   IF #_w2 THEN "DB_GlobalData".AKD.AKD1.wNewJobNumber := 4; END_IF;
   "reserve(3)":P := #_w2 AND NOT "reserve(2)";
END_REGION

REGION Network 5
   RUNG wire#powerrail
      Contact( "Clock_5Hz" )
      Coil( "xActuatorStatus" )
   END_RUNG
   // the same network as SCL:
   "xActuatorStatus" := "Clock_5Hz";
END_REGION

REGION Network 6
   #_w1 := "i_xSystemTrigger":P AND NOT "p_trig_trigg";   // rising edge
   "p_trig_trigg" := "i_xSystemTrigger":P;
   "r_eege_triger" := #_w1;
   "DB_safetyActuator".On_timer[1].TON(IN := "reserve(2)", PT := T#700ms);
END_REGION

REGION Network 7 (SCL)
   IF "r_eege_triger" THEN
       "tooglebit" := NOT "tooglebit";
   END_IF;
END_REGION

REGION Network 8
   RUNG wire#powerrail
      Contact( "DB_safetyActuator".On_timer[1].Q )
      R_Coil( "tooglebit" )
   END_RUNG
   // the same network as SCL:
   IF "DB_safetyActuator".On_timer[1].Q THEN "tooglebit" := FALSE; END_IF;
END_REGION

REGION Network 11: AKD1
   RUNG wire#powerrail
      Contact( "AKD_PNU_DATA".AKD1.PNU_userSETTINGS.xRadAKDTemp )
      Move(in := "AKD_PNU_DATA".AKD1.PNU_userSETTINGS.PNU_const.AKD_TEMP.PNU_number, out1 => "AKD_PNU_DATA".AKD1.PNU_DATA.to_PNU.iPNUnumber)
      Move(in := "AKD_PNU_DATA".AKD1.PNU_userSETTINGS.PNU_const.AKD_TEMP.PNU_subIndex, out1 => "AKD_PNU_DATA".AKD1.PNU_DATA.to_PNU.iPNUsubindex)
      Move(in := "AKD_PNU_DATA".AKD1.PNU_userSETTINGS.PNU_const.AKD_TEMP.PNU_type, out1 => "AKD_PNU_DATA".AKD1.PNU_DATA.to_PNU.wFormat)
      S_Coil( "AKD_PNU_DATA".AKD1.PNU_DATA.to_PNU.cmd.xStartRead )
      R_Coil( "AKD_PNU_DATA".AKD1.PNU_userSETTINGS.xRadAKDTemp )
   END_RUNG
   // the same network as SCL:
   IF "AKD_PNU_DATA".AKD1.PNU_userSETTINGS.xRadAKDTemp THEN
       "AKD_PNU_DATA".AKD1.PNU_DATA.to_PNU.iPNUnumber := "AKD_PNU_DATA".AKD1.PNU_userSETTINGS.PNU_const.AKD_TEMP.PNU_number;
       "AKD_PNU_DATA".AKD1.PNU_DATA.to_PNU.iPNUsubindex := "AKD_PNU_DATA".AKD1.PNU_userSETTINGS.PNU_const.AKD_TEMP.PNU_subIndex;
       "AKD_PNU_DATA".AKD1.PNU_DATA.to_PNU.wFormat := "AKD_PNU_DATA".AKD1.PNU_userSETTINGS.PNU_const.AKD_TEMP.PNU_type;
       "AKD_PNU_DATA".AKD1.PNU_DATA.to_PNU.cmd.xStartRead := TRUE;
       "AKD_PNU_DATA".AKD1.PNU_userSETTINGS.xRadAKDTemp := FALSE;
   END_IF;
END_REGION

REGION Network 12: read temperature every 0.5s
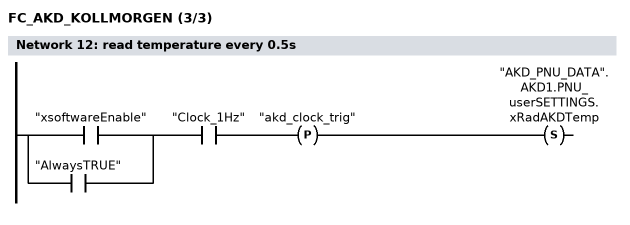
   RUNG wire#powerrail
      Contact( "xsoftwareEnable" )
      wire#w1
      Contact( "Clock_1Hz" )
      P_Trig( "akd_clock_trig" )
      S_Coil( "AKD_PNU_DATA".AKD1.PNU_userSETTINGS.xRadAKDTemp )
   END_RUNG
   RUNG wire#powerrail
      Contact( "AlwaysTRUE" )
   END_RUNG wire#w1
   // the same network as SCL:
   #_w1 := ("xsoftwareEnable" OR "AlwaysTRUE") AND "Clock_1Hz";
   #_w2 := #_w1 AND NOT "akd_clock_trig";   // rising edge
   "akd_clock_trig" := #_w1;
   IF #_w2 THEN "AKD_PNU_DATA".AKD1.PNU_userSETTINGS.xRadAKDTemp := TRUE; END_IF;
END_REGION
END_FUNCTION

FUNCTION "FC_RTD_DATA" : Void   // FC7, LAD
{ S7_Optimized_Access := 'TRUE' }
VERSION : 0.1
BEGIN

REGION Network 1
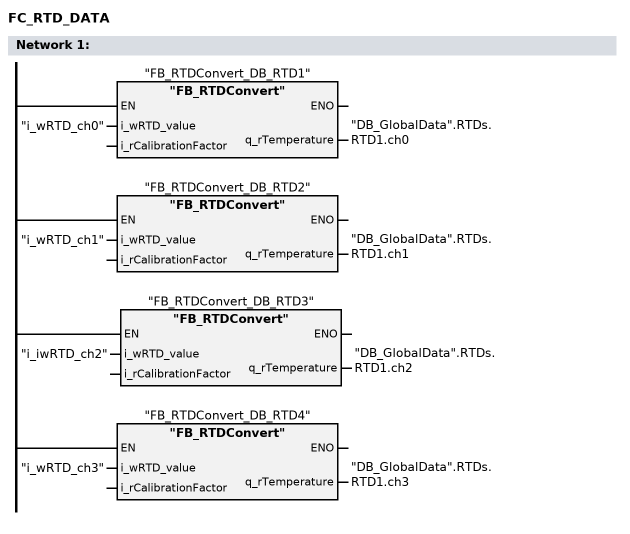
   RUNG wire#powerrail
      "FB_RTDConvert_DB_RTD1"(i_wRTD_value := "i_wRTD_ch0", i_rCalibrationFactor :=, q_rTemperature => "DB_GlobalData".RTDs.RTD1.ch0)
   END_RUNG
   RUNG wire#powerrail
      "FB_RTDConvert_DB_RTD2"(i_wRTD_value := "i_wRTD_ch1", i_rCalibrationFactor :=, q_rTemperature => "DB_GlobalData".RTDs.RTD1.ch1)
   END_RUNG
   RUNG wire#powerrail
      "FB_RTDConvert_DB_RTD3"(i_wRTD_value := "i_iwRTD_ch2", i_rCalibrationFactor :=, q_rTemperature => "DB_GlobalData".RTDs.RTD1.ch2)
   END_RUNG
   RUNG wire#powerrail
      "FB_RTDConvert_DB_RTD4"(i_wRTD_value := "i_wRTD_ch3", i_rCalibrationFactor :=, q_rTemperature => "DB_GlobalData".RTDs.RTD1.ch3)
   END_RUNG
   // the same network as SCL:
   "FB_RTDConvert_DB_RTD1"(i_wRTD_value := "i_wRTD_ch0", q_rTemperature => "DB_GlobalData".RTDs.RTD1.ch0);   // "FB_RTDConvert"
   "FB_RTDConvert_DB_RTD2"(i_wRTD_value := "i_wRTD_ch1", q_rTemperature => "DB_GlobalData".RTDs.RTD1.ch1);   // "FB_RTDConvert"
   "FB_RTDConvert_DB_RTD3"(i_wRTD_value := "i_iwRTD_ch2", q_rTemperature => "DB_GlobalData".RTDs.RTD1.ch2);   // "FB_RTDConvert"
   "FB_RTDConvert_DB_RTD4"(i_wRTD_value := "i_wRTD_ch3", q_rTemperature => "DB_GlobalData".RTDs.RTD1.ch3);   // "FB_RTDConvert"
END_REGION
END_FUNCTION

FUNCTION "FC_MQTT" : Void   // FC8, LAD
{ S7_Optimized_Access := 'TRUE' }
VERSION : 0.1
   VAR_TEMP
      globalstring : String;
      testbit : Bool;
   END_VAR
   VAR_TEMP   // added for the SCL form of the ladder/FBD networks
      _w1 : Bool;
   END_VAR
BEGIN

REGION Network 1
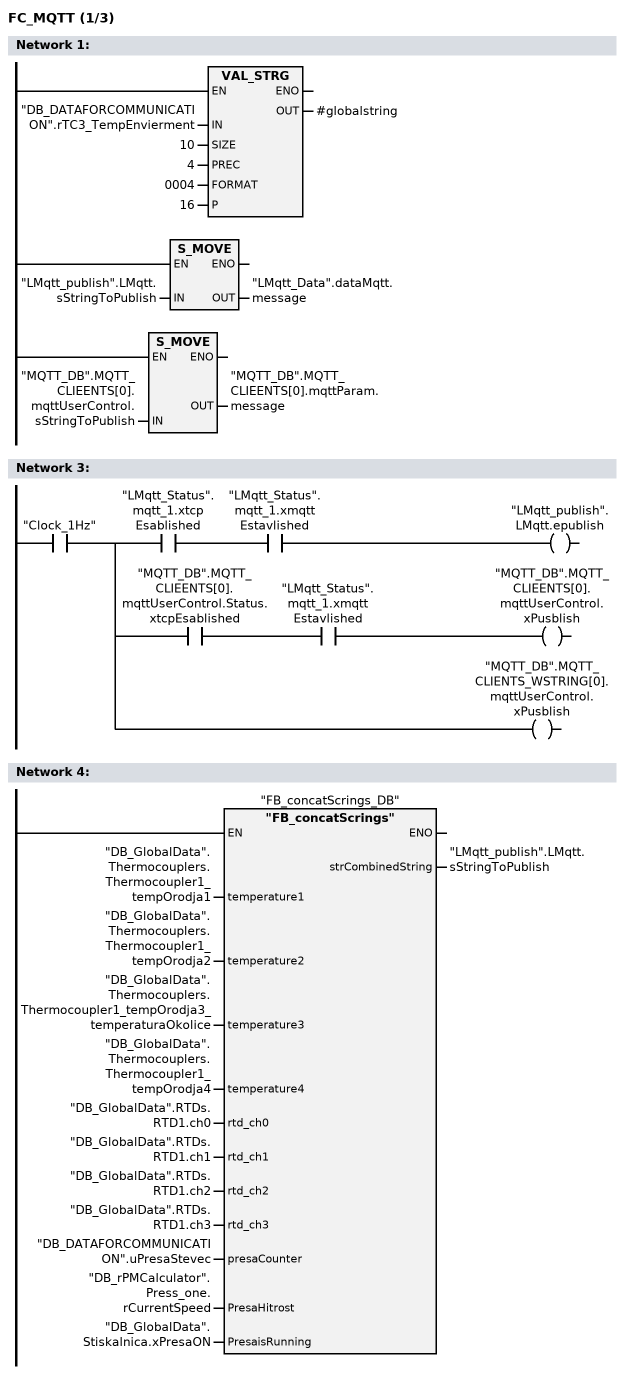
   VAL_STRG(IN := "DB_DATAFORCOMMUNICATION".rTC3_TempEnvierment,
            SIZE := 10,
            PREC := 4,
            FORMAT := 0004,
            P := 16,
            OUT => #globalstring);
   "LMqtt_Data".dataMqtt.message := "LMqtt_publish".LMqtt.sStringToPublish;
   "MQTT_DB".MQTT_CLIEENTS[0].mqttParam.message := "MQTT_DB".MQTT_CLIEENTS[0].mqttUserControl.sStringToPublish;
END_REGION

REGION Network 3
   RUNG wire#powerrail
      Contact( "Clock_1Hz" )
      wire#w1
      Contact( "LMqtt_Status".mqtt_1.xtcpEsablished )
      Contact( "LMqtt_Status".mqtt_1.xmqttEstavlished )
      Coil( "LMqtt_publish".LMqtt.epublish )
   END_RUNG
   RUNG wire#w1
      Contact( "MQTT_DB".MQTT_CLIEENTS[0].mqttUserControl.Status.xtcpEsablished )
      Contact( "LMqtt_Status".mqtt_1.xmqttEstavlished )
      Coil( "MQTT_DB".MQTT_CLIEENTS[0].mqttUserControl.xPusblish )
   END_RUNG
   RUNG wire#w1
      Coil( "MQTT_DB".MQTT_CLIENTS_WSTRING[0].mqttUserControl.xPusblish )
   END_RUNG
   // the same network as SCL:
   "LMqtt_publish".LMqtt.epublish := "Clock_1Hz" AND "LMqtt_Status".mqtt_1.xtcpEsablished AND "LMqtt_Status".mqtt_1.xmqttEstavlished;
   "MQTT_DB".MQTT_CLIEENTS[0].mqttUserControl.xPusblish := "Clock_1Hz" AND "MQTT_DB".MQTT_CLIEENTS[0].mqttUserControl.Status.xtcpEsablished AND "LMqtt_Status".mqtt_1.xmqttEstavlished;
   "MQTT_DB".MQTT_CLIENTS_WSTRING[0].mqttUserControl.xPusblish := "Clock_1Hz";
END_REGION

REGION Network 4
   RUNG wire#powerrail
      "FB_concatScrings_DB"(temperature1 := "DB_GlobalData".Thermocouplers.Thermocoupler1_tempOrodja1, temperature2 := "DB_GlobalData".Thermocouplers.Thermocoupler1_tempOrodja2, temperature3 := "DB_GlobalData".Thermocouplers.Thermocoupler1_tempOrodja3_temperaturaOkolice, temperature4 := "DB_GlobalData".Thermocouplers.Thermocoupler1_tempOrodja4, rtd_ch0 := "DB_GlobalData".RTDs.RTD1.ch0, rtd_ch1 := "DB_GlobalData".RTDs.RTD1.ch1, rtd_ch2 := "DB_GlobalData".RTDs.RTD1.ch2, rtd_ch3 := "DB_GlobalData".RTDs.RTD1.ch3, presaCounter := "DB_DATAFORCOMMUNICATION".uPresaStevec, PresaHitrost := "DB_rPMCalculator".Press_one.rCurrentSpeed, PresaisRunning := "DB_GlobalData".Stiskalnica.xPresaON, strCombinedString => "LMqtt_publish".LMqtt.sStringToPublish)
   END_RUNG
   // the same network as SCL:
   "FB_concatScrings_DB"(temperature1 := "DB_GlobalData".Thermocouplers.Thermocoupler1_tempOrodja1,   // "FB_concatScrings"
                         temperature2 := "DB_GlobalData".Thermocouplers.Thermocoupler1_tempOrodja2,
                         temperature3 := "DB_GlobalData".Thermocouplers.Thermocoupler1_tempOrodja3_temperaturaOkolice,
                         temperature4 := "DB_GlobalData".Thermocouplers.Thermocoupler1_tempOrodja4,
                         rtd_ch0 := "DB_GlobalData".RTDs.RTD1.ch0,
                         rtd_ch1 := "DB_GlobalData".RTDs.RTD1.ch1,
                         rtd_ch2 := "DB_GlobalData".RTDs.RTD1.ch2,
                         rtd_ch3 := "DB_GlobalData".RTDs.RTD1.ch3,
                         presaCounter := "DB_DATAFORCOMMUNICATION".uPresaStevec,
                         PresaHitrost := "DB_rPMCalculator".Press_one.rCurrentSpeed,
                         PresaisRunning := "DB_GlobalData".Stiskalnica.xPresaON,
                         strCombinedString => "LMqtt_publish".LMqtt.sStringToPublish);
END_REGION

REGION Network 5: MQTT publisher 1
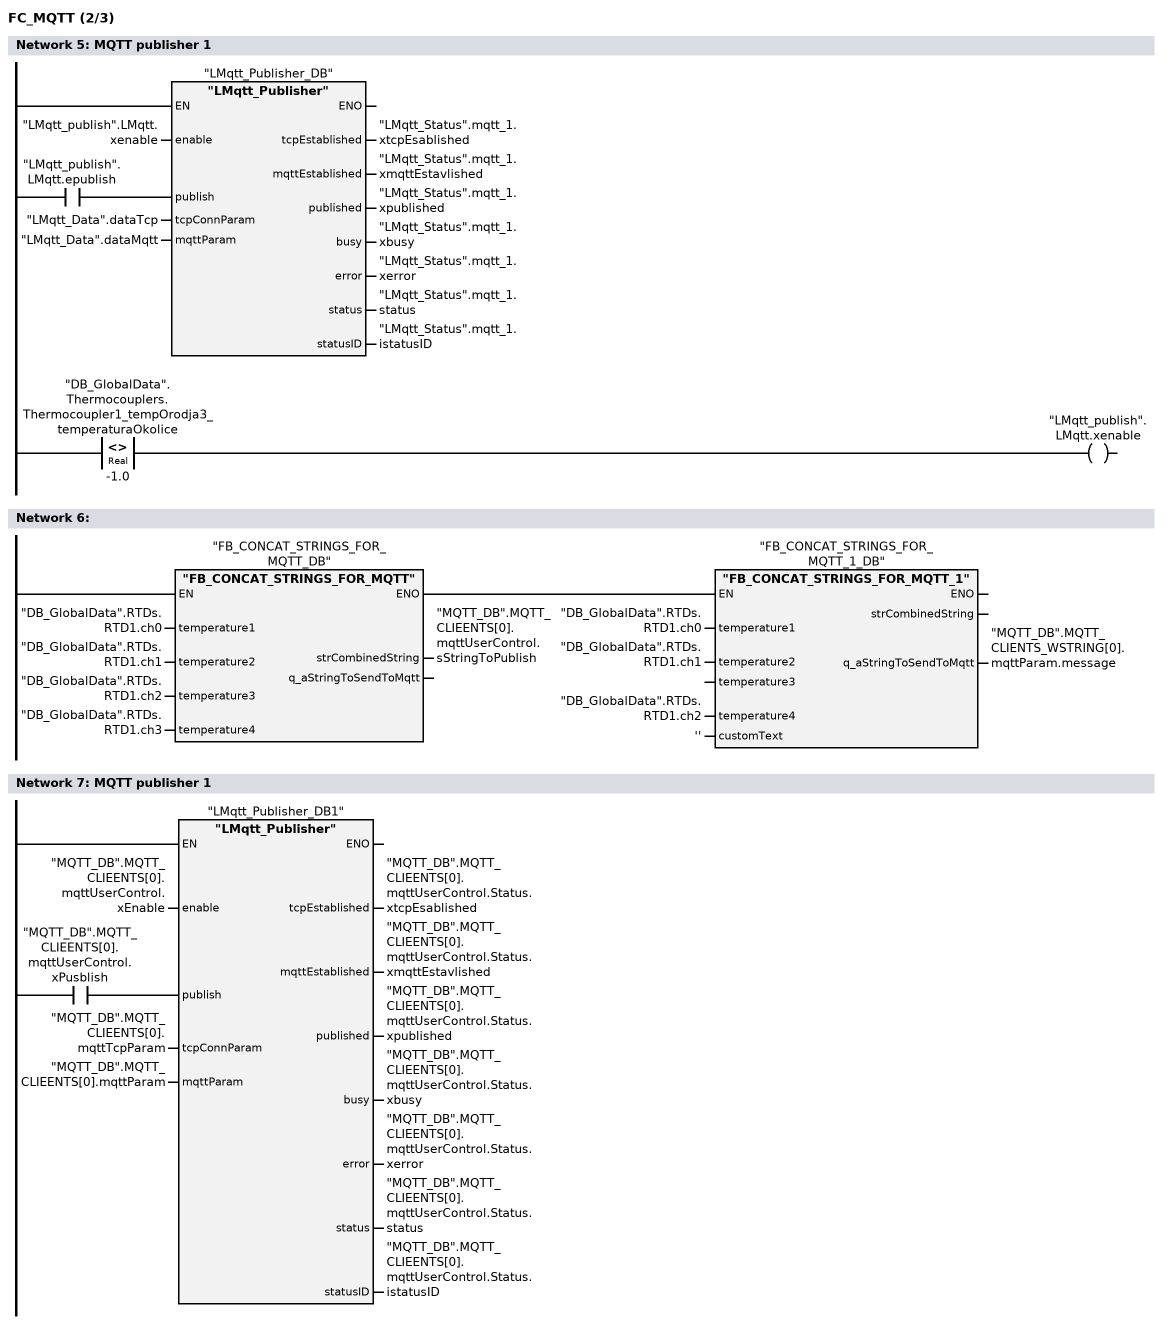
   RUNG wire#powerrail
      "LMqtt_Publisher_DB"(publish := wire#w1, enable := "LMqtt_publish".LMqtt.xenable, tcpConnParam := "LMqtt_Data".dataTcp, mqttParam := "LMqtt_Data".dataMqtt, tcpEstablished => "LMqtt_Status".mqtt_1.xtcpEsablished, mqttEstablished => "LMqtt_Status".mqtt_1.xmqttEstavlished, published => "LMqtt_Status".mqtt_1.xpublished, busy => "LMqtt_Status".mqtt_1.xbusy, error => "LMqtt_Status".mqtt_1.xerror, status => "LMqtt_Status".mqtt_1.status, statusID => "LMqtt_Status".mqtt_1.istatusID)
   END_RUNG
   RUNG wire#powerrail
      Contact( "LMqtt_publish".LMqtt.epublish )
   END_RUNG wire#w1
   RUNG wire#powerrail
      { S7_Templates := "SrcType := Real" } NE_Contact(in1 := "DB_GlobalData".Thermocouplers.Thermocoupler1_tempOrodja3_temperaturaOkolice, in2 := -1.0)
      Coil( "LMqtt_publish".LMqtt.xenable )
   END_RUNG
   // the same network as SCL:
   "LMqtt_Publisher_DB"(enable := "LMqtt_publish".LMqtt.xenable,   // "LMqtt_Publisher"
                        publish := "LMqtt_publish".LMqtt.epublish,
                        tcpConnParam := "LMqtt_Data".dataTcp,
                        mqttParam := "LMqtt_Data".dataMqtt,
                        tcpEstablished => "LMqtt_Status".mqtt_1.xtcpEsablished,
                        mqttEstablished => "LMqtt_Status".mqtt_1.xmqttEstavlished,
                        published => "LMqtt_Status".mqtt_1.xpublished,
                        busy => "LMqtt_Status".mqtt_1.xbusy,
                        error => "LMqtt_Status".mqtt_1.xerror,
                        status => "LMqtt_Status".mqtt_1.status,
                        statusID => "LMqtt_Status".mqtt_1.istatusID);
   "LMqtt_publish".LMqtt.xenable := "DB_GlobalData".Thermocouplers.Thermocoupler1_tempOrodja3_temperaturaOkolice <> (-1.0);
END_REGION

REGION Network 6
   RUNG wire#powerrail
      "FB_CONCAT_STRINGS_FOR_MQTT_DB"(temperature1 := "DB_GlobalData".RTDs.RTD1.ch0, temperature2 := "DB_GlobalData".RTDs.RTD1.ch1, temperature3 := "DB_GlobalData".RTDs.RTD1.ch2, temperature4 := "DB_GlobalData".RTDs.RTD1.ch3, strCombinedString => "MQTT_DB".MQTT_CLIEENTS[0].mqttUserControl.sStringToPublish, q_aStringToSendToMqtt =>)
      "FB_CONCAT_STRINGS_FOR_MQTT_1_DB"(temperature1 := "DB_GlobalData".RTDs.RTD1.ch0, temperature2 := "DB_GlobalData".RTDs.RTD1.ch1, temperature3 :=, temperature4 := "DB_GlobalData".RTDs.RTD1.ch2, customText := '', strCombinedString =>, q_aStringToSendToMqtt => "MQTT_DB".MQTT_CLIENTS_WSTRING[0].mqttParam.message)
   END_RUNG
   // the same network as SCL:
   "FB_CONCAT_STRINGS_FOR_MQTT_DB"(temperature1 := "DB_GlobalData".RTDs.RTD1.ch0,   // "FB_CONCAT_STRINGS_FOR_MQTT"
                           temperature2 := "DB_GlobalData".RTDs.RTD1.ch1,
                           temperature3 := "DB_GlobalData".RTDs.RTD1.ch2,
                           temperature4 := "DB_GlobalData".RTDs.RTD1.ch3,
                           strCombinedString => "MQTT_DB".MQTT_CLIEENTS[0].mqttUserControl.sStringToPublish,
                           ENO => #_w1);
   IF #_w1 THEN
       "FB_CONCAT_STRINGS_FOR_MQTT_1_DB"(temperature1 := "DB_GlobalData".RTDs.RTD1.ch0,   // "FB_CONCAT_STRINGS_FOR_MQTT_1"
                               temperature2 := "DB_GlobalData".RTDs.RTD1.ch1,
                               temperature4 := "DB_GlobalData".RTDs.RTD1.ch2,
                               customText := '',
                               q_aStringToSendToMqtt => "MQTT_DB".MQTT_CLIENTS_WSTRING[0].mqttParam.message);
   END_IF;
END_REGION

REGION Network 7: MQTT publisher 1
   RUNG wire#powerrail
      "LMqtt_Publisher_DB1"(publish := wire#w1, enable := "MQTT_DB".MQTT_CLIEENTS[0].mqttUserControl.xEnable, tcpConnParam := "MQTT_DB".MQTT_CLIEENTS[0].mqttTcpParam, mqttParam := "MQTT_DB".MQTT_CLIEENTS[0].mqttParam, tcpEstablished => "MQTT_DB".MQTT_CLIEENTS[0].mqttUserControl.Status.xtcpEsablished, mqttEstablished => "MQTT_DB".MQTT_CLIEENTS[0].mqttUserControl.Status.xmqttEstavlished, published => "MQTT_DB".MQTT_CLIEENTS[0].mqttUserControl.Status.xpublished, busy => "MQTT_DB".MQTT_CLIEENTS[0].mqttUserControl.Status.xbusy, error => "MQTT_DB".MQTT_CLIEENTS[0].mqttUserControl.Status.xerror, status => "MQTT_DB".MQTT_CLIEENTS[0].mqttUserControl.Status.status, statusID => "MQTT_DB".MQTT_CLIEENTS[0].mqttUserControl.Status.istatusID)
   END_RUNG
   RUNG wire#powerrail
      Contact( "MQTT_DB".MQTT_CLIEENTS[0].mqttUserControl.xPusblish )
   END_RUNG wire#w1
   // the same network as SCL:
   "LMqtt_Publisher_DB1"(enable := "MQTT_DB".MQTT_CLIEENTS[0].mqttUserControl.xEnable,   // "LMqtt_Publisher"
                         publish := "MQTT_DB".MQTT_CLIEENTS[0].mqttUserControl.xPusblish,
                         tcpConnParam := "MQTT_DB".MQTT_CLIEENTS[0].mqttTcpParam,
                         mqttParam := "MQTT_DB".MQTT_CLIEENTS[0].mqttParam,
                         tcpEstablished => "MQTT_DB".MQTT_CLIEENTS[0].mqttUserControl.Status.xtcpEsablished,
                         mqttEstablished => "MQTT_DB".MQTT_CLIEENTS[0].mqttUserControl.Status.xmqttEstavlished,
                         published => "MQTT_DB".MQTT_CLIEENTS[0].mqttUserControl.Status.xpublished,
                         busy => "MQTT_DB".MQTT_CLIEENTS[0].mqttUserControl.Status.xbusy,
                         error => "MQTT_DB".MQTT_CLIEENTS[0].mqttUserControl.Status.xerror,
                         status => "MQTT_DB".MQTT_CLIEENTS[0].mqttUserControl.Status.status,
                         statusID => "MQTT_DB".MQTT_CLIEENTS[0].mqttUserControl.Status.istatusID);
END_REGION

REGION Network 8: MQTT-WSTRING-TEST
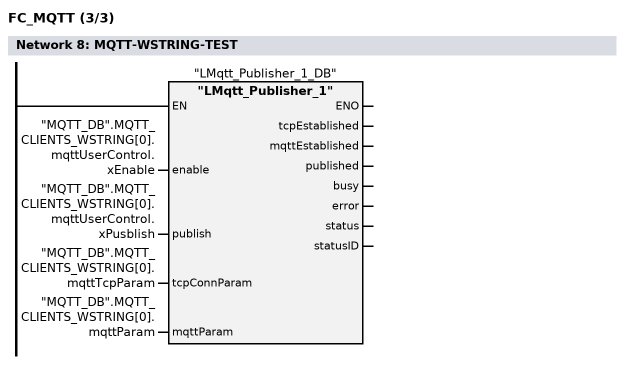
   RUNG wire#powerrail
      "LMqtt_Publisher_1_DB"(enable := "MQTT_DB".MQTT_CLIENTS_WSTRING[0].mqttUserControl.xEnable, publish := "MQTT_DB".MQTT_CLIENTS_WSTRING[0].mqttUserControl.xPusblish, tcpConnParam := "MQTT_DB".MQTT_CLIENTS_WSTRING[0].mqttTcpParam, mqttParam := "MQTT_DB".MQTT_CLIENTS_WSTRING[0].mqttParam, tcpEstablished =>, mqttEstablished =>, published =>, busy =>, error =>, status =>, statusID =>)
   END_RUNG
   // the same network as SCL:
   "LMqtt_Publisher_1_DB"(enable := "MQTT_DB".MQTT_CLIENTS_WSTRING[0].mqttUserControl.xEnable,   // "LMqtt_Publisher_1"
                          publish := "MQTT_DB".MQTT_CLIENTS_WSTRING[0].mqttUserControl.xPusblish,
                          tcpConnParam := "MQTT_DB".MQTT_CLIENTS_WSTRING[0].mqttTcpParam,
                          mqttParam := "MQTT_DB".MQTT_CLIENTS_WSTRING[0].mqttParam);
END_REGION
END_FUNCTION

FUNCTION "FC_CalculatePressRPM" : Void   // FC9, LAD
{ S7_Optimized_Access := 'TRUE' }
VERSION : 0.1
   VAR_INPUT
      i_xPulse : Bool;   // Pulse for every turn
   END_VAR
   VAR_IN_OUT
      i_iCurrentCounter : Int;
      q_iRealSPeed : Int;
   END_VAR
   VAR_TEMP
      xcalculateRPM : Bool;
      _xton : Bool;
      Temp_RPM : Real;
   END_VAR
   VAR_TEMP   // added for the SCL form of the ladder/FBD networks
      _w1 : Bool;
   END_VAR
BEGIN

REGION Network 2: 5S TIMER
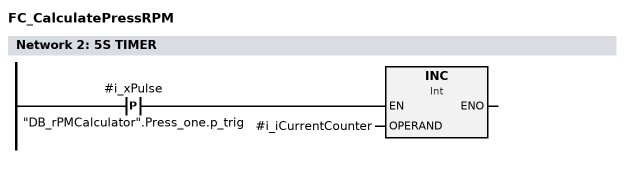
   RUNG wire#powerrail
      P_Contact(operand := #i_xPulse, bit := "DB_rPMCalculator".Press_one.p_trig)
      { S7_Templates := "DestType := Int" } Inc( #i_iCurrentCounter )
   END_RUNG
   // the same network as SCL:
   #_w1 := #i_xPulse AND NOT "DB_rPMCalculator".Press_one.p_trig;   // rising edge of #i_xPulse
   "DB_rPMCalculator".Press_one.p_trig := #i_xPulse;
   IF #_w1 THEN #i_iCurrentCounter := #i_iCurrentCounter + 1; END_IF;
END_REGION

REGION Network 3 (SCL)
   // Start 5-second timer
   "DB_rPMCalculator".Press_one.PulseTimer(IN := TRUE, PT := T#5s);



   // When 5 seconds have passed, calculate RPM
   IF "DB_rPMCalculator".Press_one.PulseTimer.Q THEN
       #q_iRealSPeed := INT_TO_REAL(#i_iCurrentCounter * 60.0) / (5.0);  // Calculate RPM
      // #q_iRealSPeed := #Temp_RPM;                      // Set the output RPM

       // Reset pulse count and timer
       #i_iCurrentCounter := 0;
       "DB_rPMCalculator".Press_one.PulseTimer(IN := FALSE,
                                               PT := T#5s);                // Reset the timer
   END_IF;
END_REGION
END_FUNCTION

FUNCTION "FC_AKD_PNU" : Void   // FC10, LAD
{ S7_Optimized_Access := 'TRUE' }
VERSION : 0.1
   VAR_INPUT
      HW_IO_telegram : Hw_Io;
   END_VAR
   VAR_IN_OUT
      AKD_PNU_v02_Instance : "AKD_PNU_v02";
      IO_DATA : "PNU_DATA";
   END_VAR
BEGIN

REGION Network 1: AKD1
   // AKD FB
   // 
   // set ID - to telegram ID of a AKD
   // 
   // 
   // # Read data from AKD PNU #
   // =================================================
   // 
   // 1. set PNU number and PNU subindex (iPNUnumber, iPNUsubindex)
   // 2. set cmd.xstartRead bit to One
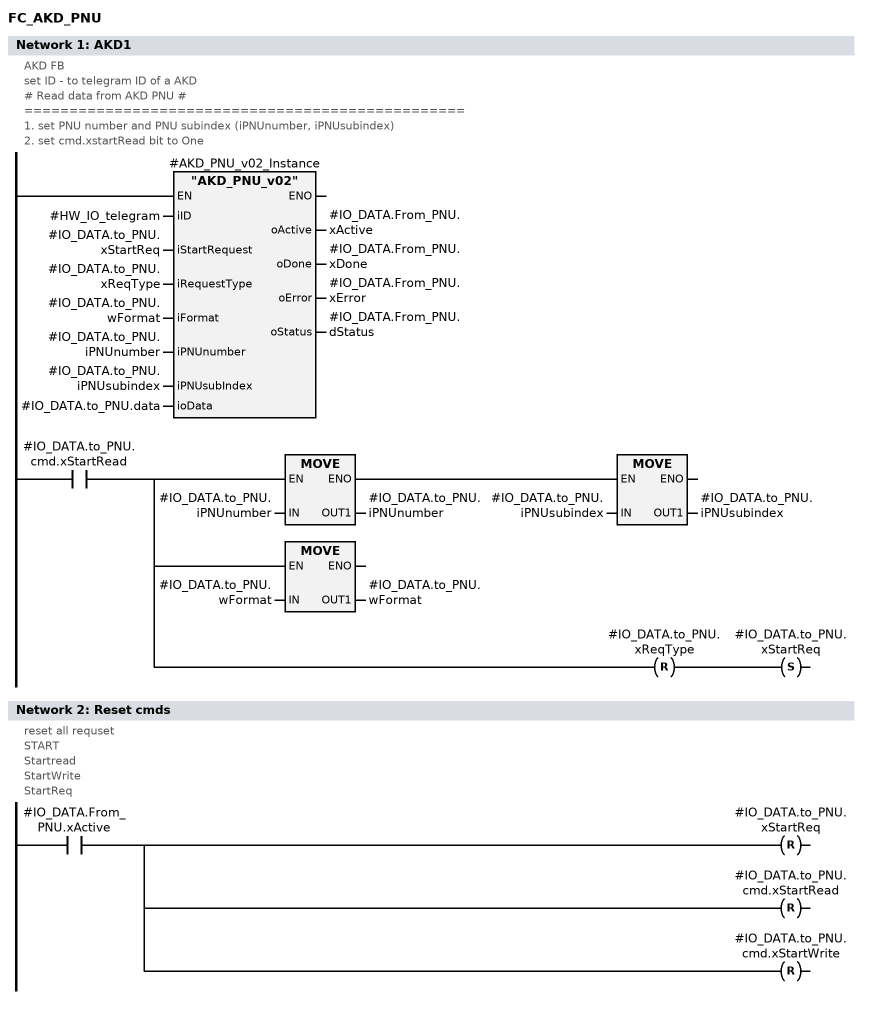
   RUNG wire#powerrail
      #AKD_PNU_v02_Instance(iID := #HW_IO_telegram, iStartRequest := #IO_DATA.to_PNU.xStartReq, iRequestType := #IO_DATA.to_PNU.xReqType, iFormat := #IO_DATA.to_PNU.wFormat, iPNUnumber := #IO_DATA.to_PNU.iPNUnumber, iPNUsubIndex := #IO_DATA.to_PNU.iPNUsubindex, ioData := #IO_DATA.to_PNU.data, oActive => #IO_DATA.From_PNU.xActive, oDone => #IO_DATA.From_PNU.xDone, oError => #IO_DATA.From_PNU.xError, oStatus => #IO_DATA.From_PNU.dStatus)
   END_RUNG
   RUNG wire#powerrail
      Contact( #IO_DATA.to_PNU.cmd.xStartRead )
      wire#w1
      Move(in := #IO_DATA.to_PNU.iPNUnumber, out1 => #IO_DATA.to_PNU.iPNUnumber)
      Move(in := #IO_DATA.to_PNU.iPNUsubindex, out1 => #IO_DATA.to_PNU.iPNUsubindex)
   END_RUNG
   RUNG wire#w1
      Move(in := #IO_DATA.to_PNU.wFormat, out1 => #IO_DATA.to_PNU.wFormat)
   END_RUNG
   RUNG wire#w1
      R_Coil( #IO_DATA.to_PNU.xReqType )
      S_Coil( #IO_DATA.to_PNU.xStartReq )
   END_RUNG
   // the same network as SCL:
   #AKD_PNU_v02_Instance(iID := #HW_IO_telegram,   // "AKD_PNU_v02"
                         iStartRequest := #IO_DATA.to_PNU.xStartReq,
                         iRequestType := #IO_DATA.to_PNU.xReqType,
                         iFormat := #IO_DATA.to_PNU.wFormat,
                         iPNUnumber := #IO_DATA.to_PNU.iPNUnumber,
                         iPNUsubIndex := #IO_DATA.to_PNU.iPNUsubindex,
                         ioData := #IO_DATA.to_PNU.data,
                         oActive => #IO_DATA.From_PNU.xActive,
                         oDone => #IO_DATA.From_PNU.xDone,
                         oError => #IO_DATA.From_PNU.xError,
                         oStatus => #IO_DATA.From_PNU.dStatus);
   IF #IO_DATA.to_PNU.cmd.xStartRead THEN
       #IO_DATA.to_PNU.iPNUnumber := #IO_DATA.to_PNU.iPNUnumber;
       #IO_DATA.to_PNU.iPNUsubindex := #IO_DATA.to_PNU.iPNUsubindex;
       #IO_DATA.to_PNU.wFormat := #IO_DATA.to_PNU.wFormat;
       #IO_DATA.to_PNU.xReqType := FALSE;
       #IO_DATA.to_PNU.xStartReq := TRUE;
   END_IF;
END_REGION

REGION Network 2: Reset cmds
   // reset all requset
   // 
   // START
   // Startread
   // StartWrite
   // StartReq
   RUNG wire#powerrail
      Contact( #IO_DATA.From_PNU.xActive )
      wire#w1
      R_Coil( #IO_DATA.to_PNU.xStartReq )
   END_RUNG
   RUNG wire#w1
      R_Coil( #IO_DATA.to_PNU.cmd.xStartRead )
   END_RUNG
   RUNG wire#w1
      R_Coil( #IO_DATA.to_PNU.cmd.xStartWrite )
   END_RUNG
   // the same network as SCL:
   IF #IO_DATA.From_PNU.xActive THEN
       #IO_DATA.to_PNU.xStartReq := FALSE;
       #IO_DATA.to_PNU.cmd.xStartRead := FALSE;
       #IO_DATA.to_PNU.cmd.xStartWrite := FALSE;
   END_IF;
END_REGION
END_FUNCTION

FUNCTION "FC_MotorControl" : Void   // FC11, LAD
{ S7_Optimized_Access := 'TRUE' }
VERSION : 0.1
   VAR_TEMP
      xM1_GoPOS2 : Bool;
      xM2_goPOS2 : Bool;
      xM3_GoPOS2 : Bool;
      xM4_GoPOS2 : Bool;
      xM5_goPOS2 : Bool;
   END_VAR
BEGIN

REGION Network 1: Cylinder CONTROL
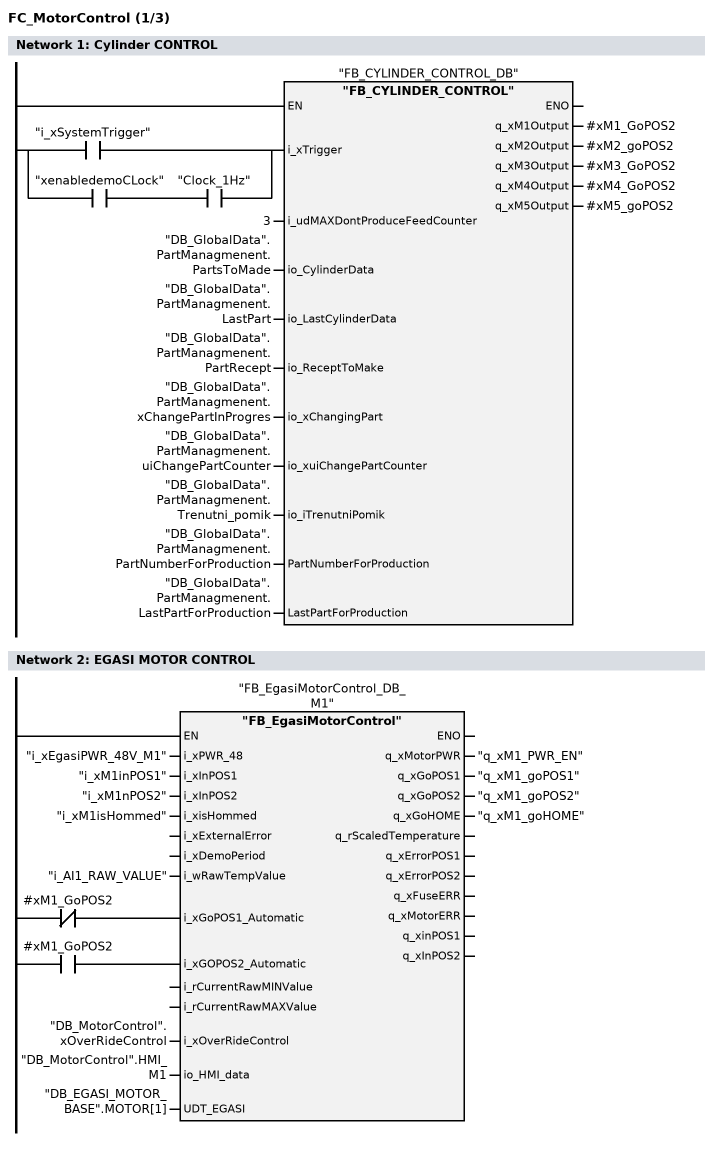
   RUNG wire#powerrail
      "FB_CYLINDER_CONTROL_DB"(i_xTrigger := wire#w1, i_udMAXDontProduceFeedCounter := 3, io_CylinderData := "DB_GlobalData".PartManagmenent.PartsToMade, io_LastCylinderData := "DB_GlobalData".PartManagmenent.LastPart, io_ReceptToMake := "DB_GlobalData".PartManagmenent.PartRecept, io_xChangingPart := "DB_GlobalData".PartManagmenent.xChangePartInProgres, io_xuiChangePartCounter := "DB_GlobalData".PartManagmenent.uiChangePartCounter, io_iTrenutniPomik := "DB_GlobalData".PartManagmenent.Trenutni_pomik, PartNumberForProduction := "DB_GlobalData".PartManagmenent.PartNumberForProduction, LastPartForProduction := "DB_GlobalData".PartManagmenent.LastPartForProduction, q_xM1Output => #xM1_GoPOS2, q_xM2Output => #xM2_goPOS2, q_xM3Output => #xM3_GoPOS2, q_xM4Output => #xM4_GoPOS2, q_xM5Output => #xM5_goPOS2)
   END_RUNG
   RUNG wire#powerrail
      Contact( "i_xSystemTrigger" )
   END_RUNG wire#w1
   RUNG wire#powerrail
      Contact( "xenabledemoCLock" )
      Contact( "Clock_1Hz" )
   END_RUNG wire#w1
   // the same network as SCL:
   "FB_CYLINDER_CONTROL_DB"(i_xTrigger := "i_xSystemTrigger" OR ("xenabledemoCLock" AND "Clock_1Hz"),   // "FB_CYLINDER_CONTROL"
                           i_udMAXDontProduceFeedCounter := 3,
                           io_CylinderData := "DB_GlobalData".PartManagmenent.PartsToMade,
                           io_LastCylinderData := "DB_GlobalData".PartManagmenent.LastPart,
                           io_ReceptToMake := "DB_GlobalData".PartManagmenent.PartRecept,
                           io_xChangingPart := "DB_GlobalData".PartManagmenent.xChangePartInProgres,
                           io_xuiChangePartCounter := "DB_GlobalData".PartManagmenent.uiChangePartCounter,
                           io_iTrenutniPomik := "DB_GlobalData".PartManagmenent.Trenutni_pomik,
                           PartNumberForProduction := "DB_GlobalData".PartManagmenent.PartNumberForProduction,
                           LastPartForProduction := "DB_GlobalData".PartManagmenent.LastPartForProduction,
                           q_xM1Output => #xM1_GoPOS2,
                           q_xM2Output => #xM2_goPOS2,
                           q_xM3Output => #xM3_GoPOS2,
                           q_xM4Output => #xM4_GoPOS2,
                           q_xM5Output => #xM5_goPOS2);
END_REGION

REGION Network 2: EGASI MOTOR CONTROL
   RUNG wire#powerrail
      "FB_EgasiMotorControl_DB_M1"(i_xGoPOS1_Automatic := wire#w1, i_xGOPOS2_Automatic := wire#w2, i_xPWR_48 := "i_xEgasiPWR_48V_M1", i_xInPOS1 := "i_xM1inPOS1", i_xInPOS2 := "i_xM1nPOS2", i_xisHommed := "i_xM1isHommed", i_xExternalError :=, i_xDemoPeriod :=, i_wRawTempValue := "i_AI1_RAW_VALUE", i_rCurrentRawMINValue :=, i_rCurrentRawMAXValue :=, i_xOverRideControl := "DB_MotorControl".xOverRideControl, io_HMI_data := "DB_MotorControl".HMI_M1, UDT_EGASI := "DB_EGASI_MOTOR_BASE".MOTOR[1], q_xMotorPWR => "q_xM1_PWR_EN", q_xGoPOS1 => "q_xM1_goPOS1", q_xGoPOS2 => "q_xM1_goPOS2", q_xGoHOME => "q_xM1_goHOME", q_rScaledTemperature =>, q_xErrorPOS1 =>, q_xErrorPOS2 =>, q_xFuseERR =>, q_xMotorERR =>, q_xinPOS1 =>, q_xInPOS2 =>)
   END_RUNG
   RUNG wire#powerrail
      I_Contact( #xM1_GoPOS2 )
   END_RUNG wire#w1
   RUNG wire#powerrail
      Contact( #xM1_GoPOS2 )
   END_RUNG wire#w2
   // the same network as SCL:
   "FB_EgasiMotorControl_DB_M1"(i_xPWR_48 := "i_xEgasiPWR_48V_M1",   // "FB_EgasiMotorControl"
                           i_xInPOS1 := "i_xM1inPOS1",
                           i_xInPOS2 := "i_xM1nPOS2",
                           i_xisHommed := "i_xM1isHommed",
                           i_wRawTempValue := "i_AI1_RAW_VALUE",
                           i_xGoPOS1_Automatic := NOT #xM1_GoPOS2,
                           i_xGOPOS2_Automatic := #xM1_GoPOS2,
                           i_xOverRideControl := "DB_MotorControl".xOverRideControl,
                           io_HMI_data := "DB_MotorControl".HMI_M1,
                           UDT_EGASI := "DB_EGASI_MOTOR_BASE".MOTOR[1],
                           q_xMotorPWR => "q_xM1_PWR_EN",
                           q_xGoPOS1 => "q_xM1_goPOS1",
                           q_xGoPOS2 => "q_xM1_goPOS2",
                           q_xGoHOME => "q_xM1_goHOME");
END_REGION

REGION Network 3
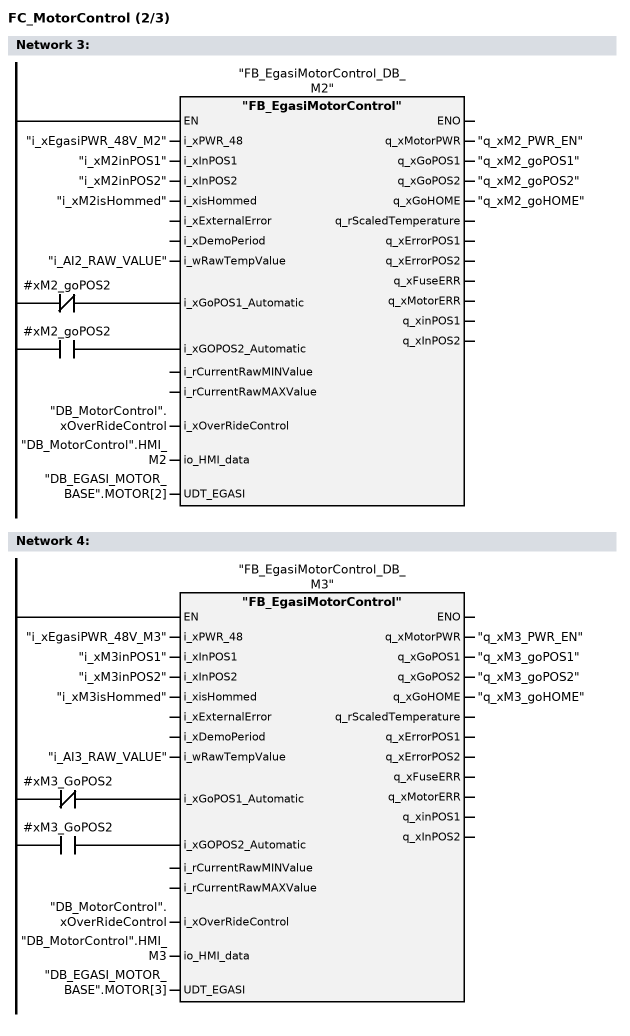
   RUNG wire#powerrail
      "FB_EgasiMotorControl_DB_M2"(i_xGoPOS1_Automatic := wire#w1, i_xGOPOS2_Automatic := wire#w2, i_xPWR_48 := "i_xEgasiPWR_48V_M2", i_xInPOS1 := "i_xM2inPOS1", i_xInPOS2 := "i_xM2inPOS2", i_xisHommed := "i_xM2isHommed", i_xExternalError :=, i_xDemoPeriod :=, i_wRawTempValue := "i_AI2_RAW_VALUE", i_rCurrentRawMINValue :=, i_rCurrentRawMAXValue :=, i_xOverRideControl := "DB_MotorControl".xOverRideControl, io_HMI_data := "DB_MotorControl".HMI_M2, UDT_EGASI := "DB_EGASI_MOTOR_BASE".MOTOR[2], q_xMotorPWR => "q_xM2_PWR_EN", q_xGoPOS1 => "q_xM2_goPOS1", q_xGoPOS2 => "q_xM2_goPOS2", q_xGoHOME => "q_xM2_goHOME", q_rScaledTemperature =>, q_xErrorPOS1 =>, q_xErrorPOS2 =>, q_xFuseERR =>, q_xMotorERR =>, q_xinPOS1 =>, q_xInPOS2 =>)
   END_RUNG
   RUNG wire#powerrail
      I_Contact( #xM2_goPOS2 )
   END_RUNG wire#w1
   RUNG wire#powerrail
      Contact( #xM2_goPOS2 )
   END_RUNG wire#w2
   // the same network as SCL:
   "FB_EgasiMotorControl_DB_M2"(i_xPWR_48 := "i_xEgasiPWR_48V_M2",   // "FB_EgasiMotorControl"
                           i_xInPOS1 := "i_xM2inPOS1",
                           i_xInPOS2 := "i_xM2inPOS2",
                           i_xisHommed := "i_xM2isHommed",
                           i_wRawTempValue := "i_AI2_RAW_VALUE",
                           i_xGoPOS1_Automatic := NOT #xM2_goPOS2,
                           i_xGOPOS2_Automatic := #xM2_goPOS2,
                           i_xOverRideControl := "DB_MotorControl".xOverRideControl,
                           io_HMI_data := "DB_MotorControl".HMI_M2,
                           UDT_EGASI := "DB_EGASI_MOTOR_BASE".MOTOR[2],
                           q_xMotorPWR => "q_xM2_PWR_EN",
                           q_xGoPOS1 => "q_xM2_goPOS1",
                           q_xGoPOS2 => "q_xM2_goPOS2",
                           q_xGoHOME => "q_xM2_goHOME");
END_REGION

REGION Network 4
   RUNG wire#powerrail
      "FB_EgasiMotorControl_DB_M3"(i_xGoPOS1_Automatic := wire#w1, i_xGOPOS2_Automatic := wire#w2, i_xPWR_48 := "i_xEgasiPWR_48V_M3", i_xInPOS1 := "i_xM3inPOS1", i_xInPOS2 := "i_xM3inPOS2", i_xisHommed := "i_xM3isHommed", i_xExternalError :=, i_xDemoPeriod :=, i_wRawTempValue := "i_AI3_RAW_VALUE", i_rCurrentRawMINValue :=, i_rCurrentRawMAXValue :=, i_xOverRideControl := "DB_MotorControl".xOverRideControl, io_HMI_data := "DB_MotorControl".HMI_M3, UDT_EGASI := "DB_EGASI_MOTOR_BASE".MOTOR[3], q_xMotorPWR => "q_xM3_PWR_EN", q_xGoPOS1 => "q_xM3_goPOS1", q_xGoPOS2 => "q_xM3_goPOS2", q_xGoHOME => "q_xM3_goHOME", q_rScaledTemperature =>, q_xErrorPOS1 =>, q_xErrorPOS2 =>, q_xFuseERR =>, q_xMotorERR =>, q_xinPOS1 =>, q_xInPOS2 =>)
   END_RUNG
   RUNG wire#powerrail
      I_Contact( #xM3_GoPOS2 )
   END_RUNG wire#w1
   RUNG wire#powerrail
      Contact( #xM3_GoPOS2 )
   END_RUNG wire#w2
   // the same network as SCL:
   "FB_EgasiMotorControl_DB_M3"(i_xPWR_48 := "i_xEgasiPWR_48V_M3",   // "FB_EgasiMotorControl"
                           i_xInPOS1 := "i_xM3inPOS1",
                           i_xInPOS2 := "i_xM3inPOS2",
                           i_xisHommed := "i_xM3isHommed",
                           i_wRawTempValue := "i_AI3_RAW_VALUE",
                           i_xGoPOS1_Automatic := NOT #xM3_GoPOS2,
                           i_xGOPOS2_Automatic := #xM3_GoPOS2,
                           i_xOverRideControl := "DB_MotorControl".xOverRideControl,
                           io_HMI_data := "DB_MotorControl".HMI_M3,
                           UDT_EGASI := "DB_EGASI_MOTOR_BASE".MOTOR[3],
                           q_xMotorPWR => "q_xM3_PWR_EN",
                           q_xGoPOS1 => "q_xM3_goPOS1",
                           q_xGoPOS2 => "q_xM3_goPOS2",
                           q_xGoHOME => "q_xM3_goHOME");
END_REGION

REGION Network 5
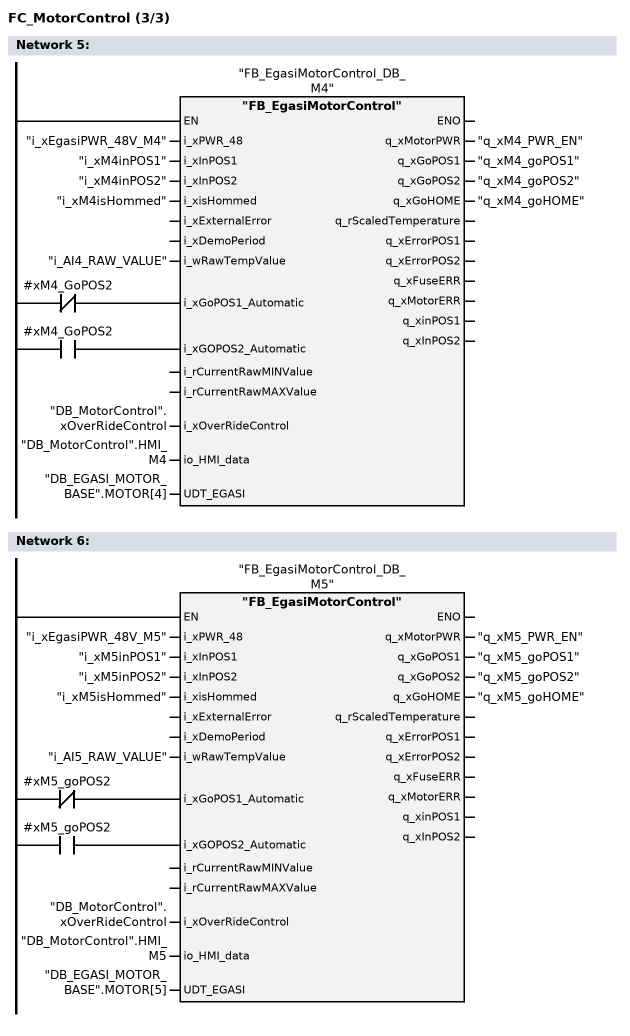
   RUNG wire#powerrail
      "FB_EgasiMotorControl_DB_M4"(i_xGoPOS1_Automatic := wire#w1, i_xGOPOS2_Automatic := wire#w2, i_xPWR_48 := "i_xEgasiPWR_48V_M4", i_xInPOS1 := "i_xM4inPOS1", i_xInPOS2 := "i_xM4inPOS2", i_xisHommed := "i_xM4isHommed", i_xExternalError :=, i_xDemoPeriod :=, i_wRawTempValue := "i_AI4_RAW_VALUE", i_rCurrentRawMINValue :=, i_rCurrentRawMAXValue :=, i_xOverRideControl := "DB_MotorControl".xOverRideControl, io_HMI_data := "DB_MotorControl".HMI_M4, UDT_EGASI := "DB_EGASI_MOTOR_BASE".MOTOR[4], q_xMotorPWR => "q_xM4_PWR_EN", q_xGoPOS1 => "q_xM4_goPOS1", q_xGoPOS2 => "q_xM4_goPOS2", q_xGoHOME => "q_xM4_goHOME", q_rScaledTemperature =>, q_xErrorPOS1 =>, q_xErrorPOS2 =>, q_xFuseERR =>, q_xMotorERR =>, q_xinPOS1 =>, q_xInPOS2 =>)
   END_RUNG
   RUNG wire#powerrail
      I_Contact( #xM4_GoPOS2 )
   END_RUNG wire#w1
   RUNG wire#powerrail
      Contact( #xM4_GoPOS2 )
   END_RUNG wire#w2
   // the same network as SCL:
   "FB_EgasiMotorControl_DB_M4"(i_xPWR_48 := "i_xEgasiPWR_48V_M4",   // "FB_EgasiMotorControl"
                           i_xInPOS1 := "i_xM4inPOS1",
                           i_xInPOS2 := "i_xM4inPOS2",
                           i_xisHommed := "i_xM4isHommed",
                           i_wRawTempValue := "i_AI4_RAW_VALUE",
                           i_xGoPOS1_Automatic := NOT #xM4_GoPOS2,
                           i_xGOPOS2_Automatic := #xM4_GoPOS2,
                           i_xOverRideControl := "DB_MotorControl".xOverRideControl,
                           io_HMI_data := "DB_MotorControl".HMI_M4,
                           UDT_EGASI := "DB_EGASI_MOTOR_BASE".MOTOR[4],
                           q_xMotorPWR => "q_xM4_PWR_EN",
                           q_xGoPOS1 => "q_xM4_goPOS1",
                           q_xGoPOS2 => "q_xM4_goPOS2",
                           q_xGoHOME => "q_xM4_goHOME");
END_REGION

REGION Network 6
   RUNG wire#powerrail
      "FB_EgasiMotorControl_DB_M5"(i_xGoPOS1_Automatic := wire#w1, i_xGOPOS2_Automatic := wire#w2, i_xPWR_48 := "i_xEgasiPWR_48V_M5", i_xInPOS1 := "i_xM5inPOS1", i_xInPOS2 := "i_xM5inPOS2", i_xisHommed := "i_xM5isHommed", i_xExternalError :=, i_xDemoPeriod :=, i_wRawTempValue := "i_AI5_RAW_VALUE", i_rCurrentRawMINValue :=, i_rCurrentRawMAXValue :=, i_xOverRideControl := "DB_MotorControl".xOverRideControl, io_HMI_data := "DB_MotorControl".HMI_M5, UDT_EGASI := "DB_EGASI_MOTOR_BASE".MOTOR[5], q_xMotorPWR => "q_xM5_PWR_EN", q_xGoPOS1 => "q_xM5_goPOS1", q_xGoPOS2 => "q_xM5_goPOS2", q_xGoHOME => "q_xM5_goHOME", q_rScaledTemperature =>, q_xErrorPOS1 =>, q_xErrorPOS2 =>, q_xFuseERR =>, q_xMotorERR =>, q_xinPOS1 =>, q_xInPOS2 =>)
   END_RUNG
   RUNG wire#powerrail
      I_Contact( #xM5_goPOS2 )
   END_RUNG wire#w1
   RUNG wire#powerrail
      Contact( #xM5_goPOS2 )
   END_RUNG wire#w2
   // the same network as SCL:
   "FB_EgasiMotorControl_DB_M5"(i_xPWR_48 := "i_xEgasiPWR_48V_M5",   // "FB_EgasiMotorControl"
                           i_xInPOS1 := "i_xM5inPOS1",
                           i_xInPOS2 := "i_xM5inPOS2",
                           i_xisHommed := "i_xM5isHommed",
                           i_wRawTempValue := "i_AI5_RAW_VALUE",
                           i_xGoPOS1_Automatic := NOT #xM5_goPOS2,
                           i_xGOPOS2_Automatic := #xM5_goPOS2,
                           i_xOverRideControl := "DB_MotorControl".xOverRideControl,
                           io_HMI_data := "DB_MotorControl".HMI_M5,
                           UDT_EGASI := "DB_EGASI_MOTOR_BASE".MOTOR[5],
                           q_xMotorPWR => "q_xM5_PWR_EN",
                           q_xGoPOS1 => "q_xM5_goPOS1",
                           q_xGoPOS2 => "q_xM5_goPOS2",
                           q_xGoHOME => "q_xM5_goHOME");
END_REGION
END_FUNCTION

FUNCTION "FC_PARTMANAGE" : Void   // FC12, LAD
{ S7_Optimized_Access := 'TRUE' }
VERSION : 0.1
   VAR_TEMP   // added for the SCL form of the ladder/FBD networks
      _w1 : Bool;
   END_VAR
BEGIN

REGION Network 2: COPY DATA FROM BASE TO DB for Cylinder control
